// Mitsubishi GX Works2 project: 701125增加出库   PLC: Q10UDEH (continued)
IF iStep=3 AND ConveyorMotor.xSizeDeficientDetect AND (NOT ConveyorMotor.xCCWPresent OR NOT ConveyorMotor.xCWPresent)  THEN
	   ConveyorMotor.xOverWidthAlarm:=1;
	    iStep:=0;               
END_IF;
(*//总报警*)
ConveyorMotor.xError:=ConveyorMotor.xLimitAlarrm
                                              OR ConveyorMotor.xNotArriveAlarm
                                              OR ConveyorMotor.xUnloadAlarm                                             
                                              OR ConveyorMotor.xOverWidthAlarm;

(*//状态输出*)(*状态显示，容易造成指针容量不足*)
IF ConveyorMotor.xEmpty AND NOT ConveyorMotor.xBusy THEN
	m_wStateWord:=0;
END_IF;
IF ConveyorMotor.xEmpty=0 THEN
		m_wStateWord:=1;
END_IF;
IF ConveyorMotor.xBusy THEN
		m_wStateWord:=2;
END_IF;
IF ConveyorMotor.xLimitAlarrm THEN
		m_wStateWord:=3;
END_IF;
IF ConveyorMotor.xOverWidthAlarm THEN
		m_wStateWord:=4;
END_IF;
IF ConveyorMotor.xNotArriveAlarm THEN	
		m_wStateWord:=5;
END_IF;
IF ConveyorMotor.xUnloadAlarm THEN
		m_wStateWord:=6;	
END_IF;
(*选择本线体后，将状态赋值给全局变量进行显示*)
IF ConveyorMotor.iDeviceID=g_iDeviceIDSelect THEN
	g_iConveyorStatus:=m_wStateWord;
END_IF;
END_FUNCTION_BLOCK

FUNCTION_BLOCK DivideFolder
VAR_IN_OUT
  FolderIO : FolderIO;
  FolderConveyorIO : ConveyorIO;
END_VAR
VAR
  iFolderCount : INT;
  m_xInitial : BOOL;
  istep : INT;
  m_TONLoadDelay : TON;  (* 上料完成延时 *)
  m_xLoadDelay : BOOL;  (* 上料完成延时 *)
  m_tLoadDelay : TIME;  (* 上料完成延时 *)
  m_TONUpCylinderError : TON;
  m_tUpCylinderError : TIME;
  m_TONDownCylinderError : TON;
  m_tDownCylinderError : TIME;
  m_TONGrabCylinderError : TON;
  m_tGrabCylinderError : TIME;
END_VAR
VAR_INPUT
  i_xAuto : BOOL;  (* 自动 *)
END_VAR
(*拆盘机*)
(*Mr.Li修改2018.11.19调试*)
(*初始化*)
IF NOT m_xInitial  THEN
	FolderIO.i_iFloor:=3;
	 iFolderCount:=3;
	 	FolderIO.i_tSetOvertime:=T#5S;
		m_xInitial:=1;
END_IF;
(*自动*)
IF i_xAuto THEN
	FolderIO.o_xEntryPermit:=iFolderCount=3 AND FolderConveyorIO.xEmpty;(*线体状态为空且拆盘初始数量为3，才准上料*)
	m_TONLoadDelay(IN:= NOT FolderConveyorIO.xEmpty,
											PT:= T#100MS,
											Q:=m_xLoadDelay,
											ET:=m_tLoadDelay);

	CASE istep OF
		0:(*各种初始化*)
			FolderConveyorIO.xLoad:=0;
			FolderConveyorIO.xUnload:=0;
			FolderConveyorIO.xPutInto:=0;
			IF FolderConveyorIO.xEmpty THEN(*空的情况，0时上料，其他走流程*)
				IF iFolderCount=FolderIO.i_iFloor   THEN
					istep:=1; 					
				ELSE
					istep:=5;
				END_IF;	
			END_IF;		
			IF m_xLoadDelay THEN
				 IF FolderIO.i_xCylinderDownRetractDetect AND FolderIO.i_xCylinderUpRetractDetect THEN
					istep:=2;(*如果在1层，则顶起，需人为判断是否在指定位置，否则有翻框的危险*)
				ELSE
				 	istep:=3;(*如果有料不在1层，则抓紧，然后跳到第4步判断是否是叠盘，不是就放行*)
				 END_IF;
			END_IF;
		1:(*上料*)
			IF FolderIO.o_xEntryPermit THEN
				FolderConveyorIO.xLoad:=FolderIO.i_FrontConveyorNextRun;
			ELSE
				FolderConveyorIO.xLoad:=0;
			END_IF;(*有料等延时*)	
			IF m_xLoadDelay THEN
				iFolderCount:=FolderIO.i_iFloor;
				istep:=2;(**拆盘机顶起步骤*)
			END_IF;	
		2:(*上升至2层位置*)
				FolderIO.o_xCylinderDownRetract:=0;
				FolderIO.o_xCylinderDownExtend:=1;
				FolderIO.o_xCylinderUpRetract:=0;
				IF FolderIO.i_xCylinderDownExtendDetect   THEN
				istep:=3;
				END_IF;
		3:	(*夹紧夹爪*)
			IF FolderIO.i_xCylinderDownExtendDetect THEN
				FolderIO.o_xCylinderGrabExtend:=1;
				FolderIO.o_xCylinderGrabRetract:=0;
			END_IF;
			IF FolderIO.i_xCylinderGrabExtendDetect THEN
				istep:=4;
			END_IF;	
		4:(*再下降到1层，然后放行，在该位置判断是不是最后一次*)
				FolderIO.o_xCylinderUpRetract:=1;
				FolderIO.o_xCylinderUpExtend:=0;
				FolderIO.o_xCylinderDownRetract:=1;
				FolderIO.o_xCylinderDownExtend:=0;
				IF FolderIO.i_xCylinderDownRetractDetect AND FolderIO.i_xCylinderUpRetractDetect AND FolderIO.o_xExitPremit THEN
				FolderConveyorIO.xPutInto:=1;
				FolderConveyorIO.xUnload:=FolderIO.o_xExitPremit;
				ELSIF NOT FolderIO.i_xTrayDetect AND NOT FolderConveyorIO.xEmpty AND FolderIO.o_xExitPremit THEN 
						FolderConveyorIO.xUnload:=FolderIO.o_xExitPremit;
				ELSE 
					FolderConveyorIO.xPutInto:=0;
				FolderConveyorIO.xUnload:=0;
				END_IF;
					IF FolderIO.i_xCylinderDownRetractDetect AND FolderIO.i_xCylinderUpRetractDetect AND
						  FolderIO.i_xTrayDetect  AND  iFolderCount>0  AND ldp(TRUE,NOT  FolderConveyorIO.xUnload) THEN
						iFolderCount:=FolderIO.i_iFloor-1;					
					istep:=5;
					ELSIF  FolderIO.i_xCylinderDownRetractDetect AND FolderIO.i_xCylinderUpRetractDetect  AND 
						 NOT FolderIO.i_xTrayDetect   AND  FolderConveyorIO.xEmpty THEN 
						 	istep:=7;
					END_IF;

		5:(*上升到3层*)
			FolderIO.o_xCylinderUpRetract:=0;
			FolderIO.o_xCylinderUpExtend:=1;
			FolderIO.o_xCylinderDownRetract:=0;
			IF  FolderIO.i_xCylinderUpExtendDetect THEN
				istep:=6;
			END_IF;		
		6:(*松开并下降*)
			FolderIO.i_iFloor:=iFolderCount;
			IF  FolderIO.i_xCylinderUpExtendDetect  THEN
				FolderIO.o_xCylinderGrabExtend:=0;
				FolderIO.o_xCylinderGrabRetract:=1;
				IF FolderIO.i_xCylinderGrabRetractDetect THEN
					FolderIO.o_xCylinderUpRetract:=1;
					FolderIO.o_xCylinderUpExtend:=0;
					FolderIO.o_xCylinderDownRetract:=1;
					FolderIO.o_xCylinderDownExtend:=0;
				END_IF;		
			END_IF;	
			IF   FolderIO.i_xCylinderUpRetractDetect  AND FolderIO.i_xCylinderDownRetractDetect  THEN
				istep:=2;
			ELSIF iFolderCount=0 THEN 
				istep:=7;
			ELSIF  NOT FolderIO.i_xTrayDetect  THEN 
				istep:=4;
			END_IF;	
			
		7:(*恢复初始状态*)	
			FolderIO.o_xCylinderDownRetract:=1;
			FolderIO.o_xCylinderUpRetract:=1;
			FolderIO.o_xCylinderDownExtend:=0;
			FolderIO.o_xCylinderUpExtend:=0;
			FolderIO.o_xCylinderGrabExtend:=0;
			FolderIO.o_xCylinderGrabRetract:=1;
			iFolderCount:=3;
			FolderIO.i_iFloor:=3;
			IF FolderIO.i_xCylinderDownRetractDetect  AND FolderIO.i_xCylinderUpRetractDetect THEN 
			istep:=0;
			END_IF;
		END_CASE;
END_IF;(*g_xAuto那个*)	
(*手动控制气缸动作*)
		IF NOT i_xAuto THEN
			FolderIO.o_xCylinderGrabExtend:=	FolderIO.i_xCylinderGrabExtendButton;	
			FolderIO.o_xCylinderGrabRetract:=	FolderIO.i_xCylinderGrabRetractButton;	
			FolderIO.o_xCylinderUpExtend:=		FolderIO.i_xCylinderUpExtendButton;	
			FolderIO.o_xCylinderUpRetract:=		FolderIO.i_xCylinderUpRetractButton;	
			FolderIO.o_xCylinderDownExtend:=	FolderIO.i_xCylinderDownExtendButton;	
			FolderIO.o_xCylinderDownRetract:=	FolderIO.i_xCylinderDownRetractButton;		
		END_IF;
		
		(*气缸超时未到达报警，可能是没气儿漏气，也可能是开关坏了，或者气缸被卡住了*)
		m_TONGrabCylinderError(IN:= (FolderIO.o_xCylinderGrabExtend AND NOT FolderIO.i_xCylinderGrabExtendDetect) 
																OR  (FolderIO.o_xCylinderGrabRetract AND NOT FolderIO.i_xCylinderGrabRetractDetect) ,
															PT:= FolderIO.i_tSetOvertime ,Q:= FolderIO.o_xGrabCylinderError,ET:= m_tGrabCylinderError);
		m_TONDownCylinderError(IN:= (FolderIO.o_xCylinderDownExtend AND NOT FolderIO.i_xCylinderDownExtendDetect) 
																OR  (FolderIO.o_xCylinderDownRetract AND NOT FolderIO.i_xCylinderDownRetractDetect) ,
															PT:= FolderIO.i_tSetOvertime ,Q:= FolderIO.o_xDownCylinderError,ET:= m_tDownCylinderError);
		m_TONUpCylinderError(IN:= (FolderIO.o_xCylinderUpExtend AND NOT FolderIO.i_xCylinderUpExtendDetect) 
																OR  (FolderIO.o_xCylinderUpRetract AND NOT FolderIO.i_xCylinderUpRetractDetect) ,
															PT:= FolderIO.i_tSetOvertime ,Q:= FolderIO.o_xUpCylinderError,ET:= m_tUpCylinderError);
END_FUNCTION_BLOCK

FUNCTION_BLOCK FanucRobot
VAR_IN_OUT
  FanucRobotIO : FanucRobotIO;
END_VAR
VAR
  m_iSNO : INT;
  m_xPNSPass : BOOL;  (* 收到程序号 *)
  m_tonStartDelay : TON;  (* 启动延时 *)
  m_xStartDelay : BOOL;
  m_tStartDelayCurrentTime : TIME;
END_VAR
(***********************************************************
发那科机器人自动启动程序


***********************************************************)

(*无自动状态，示教盒处于本地状态，把各标志位复位*)
IF FanucRobotIO.i_xTPENBL AND NOT g_xAuto THEN
	FanucRobotIO.o_xPNSTROBE:=0;
	FanucRobotIO.o_xCSTOPI:=0;
	FanucRobotIO.o_xPROD_START:=0;
	FanucRobotIO.o_xRESET:=0;
END_IF;
(*远程模式*)
IF g_xAuto THEN
	FanucRobotIO.o_xREMOTE:=1;
	ELSE
	FanucRobotIO.o_xREMOTE:=0;
END_IF;
(*程序启动后复位启动标志位*)
IF FanucRobotIO.i_xPROG_RUN AND FanucRobotIO.i_xBUSY THEN
	FanucRobotIO.i_xCommandStart:=0;
END_IF;
(*示教盒旋清除报警*)
IF ldf(TRUE,FanucRobotIO.i_xTPENBL)THEN
	FanucRobotIO.o_xRESET:=1;
	FanucRobotIO.o_xCSTOPI:=1;
END_IF;
(*启动程序号条件*)
IF FanucRobotIO.i_xSYSRDY 
	AND FanucRobotIO.i_xCMDENBL
	AND FanucRobotIO.i_xCommandStart
	AND NOT FanucRobotIO.i_xPROG_RUN 
	AND NOT FanucRobotIO.i_xBUSY THEN
	FanucRobotIO.o_xRESET:=0;
	FanucRobotIO.o_xCSTOPI:=0;
	IF FanucRobotIO.i_iMotionNumber <> 0 (*只要动作编号不为0，就给他信号*)
		AND NOT FanucRobotIO.o_xPNSTROBE THEN
		FanucRobotIO.o_xPNSTROBE:=1;
		FanucRobotIO.o_xPROD_START:=1;
		FanucRobotIO.o_iPNS:=FanucRobotIO.i_iMotionNumber;(*并把任务号传给他*)
	END_IF;
	(*程序号校验*)
	IF FanucRobotIO.i_xSNACK THEN(*数据传回之后再校验*)
		m_iSNO:=BITARR_TO_INT(FanucRobotIO.i_arrxSNO[0] , 8 );
		IF m_iSNO=FanucRobotIO.o_iPNS THEN
			m_xPNSPass:=1;(*校验成功,等100MS复位Start信号*)
			FanucRobotIO.o_xPNSTROBE:=0;
		ELSE
			FanucRobotIO.o_xPNSFailed:=1;(*校验失败*)
			FanucRobotIO.o_xPROD_START:=0;(*立刻复位，不生成任务*)
		END_IF;
	END_IF;
END_IF;
m_tonStartDelay(IN:= m_xPNSPass ,PT:= T#100ms ,Q:= m_xStartDelay ,ET:=m_tStartDelayCurrentTime );
IF m_xStartDelay THEN
	FanucRobotIO.o_xPROD_START:=0;
	FanucRobotIO.i_xCommandStart:=0;
	m_xPNSPass:=0;
END_IF;
END_FUNCTION_BLOCK

FUNCTION_BLOCK Folder
VAR_IN_OUT
  FolderIO : FolderIO;
END_VAR
VAR
  m_xInitial : BOOL;
END_VAR
VAR_IN_OUT
  FolderConveyorIO : ConveyorIO;
END_VAR
VAR
  iFolderCount : INT;
  istep : INT;
  m_TONLoadDelay : TON;  (* 上料完成延时 *)
  m_xLoadDelay : BOOL;  (* 上料完成延时 *)
  m_tLoadDelay : TIME;  (* 上料完成延时 *)
  m_TONUpCylinderError : TON;
  m_tUpCylinderError : TIME;
  m_TONDownCylinderError : TON;
  m_tDownCylinderError : TIME;
  m_TONGrabCylinderError : TON;
  m_tGrabCylinderError : TIME;
END_VAR
VAR_INPUT
  i_xAuto : BOOL;  (* 自动 *)
  i_xManual : BOOL;  (* 手动 *)
END_VAR
(*叠盘机*)
(*sb刘写的*)
(*初始化*)
(*18/11/17 YAOBO更改*)
(*增加允许下料信号o_xExitPrimit，码垛完成后给允许下料第7步给出*)
IF NOT m_xInitial THEN
	FolderIO.i_iFloor:=3;
	FolderIO.i_tSetOvertime:=T#5S;
	
	m_xInitial:=1;
END_IF;
(*自动*)
FolderIO.o_xEntryPermit:=FolderConveyorIO.xEmpty;(*叠盘机的话，只要空了，就允许上料，拆盘则是拆完才允许*)
IF i_xAuto THEN
				m_TONLoadDelay(IN:= NOT FolderConveyorIO.xEmpty,
													PT:= T#100MS,
													Q:=m_xLoadDelay,
													ET:=m_tLoadDelay);
	CASE istep OF
		0:(*各种初始化*)
			FolderConveyorIO.xLoad:=0;
			FolderConveyorIO.xUnload:=0;
			FolderConveyorIO.xPutInto:=0;
			FolderIo.o_xExitPremit:=0;	
			IF (*0 AND*)  FolderConveyorIO.xEmpty THEN
				istep:=1;(*空着就去1上料*)
			END_IF;	
			IF 0 AND    m_xLoadDelay  THEN(*if 有料*)
				IF  FolderIO.i_xCylinderDownExtendDetect  AND FolderIO.i_xCylinderUpExtendDetect  THEN(*if 在下层*)
					IF iFolderCount=FolderIO.i_iFloor THEN(*if 是最后一次*)
						istep:=7;
					ELSE(*不是最后一次去5，是就去7*)
						istep:=5;
					END_IF;(*if 是最后一次*)	
				ELSE(*不在下层去2*)
				istep:=2;
				END_IF;	(*if 在下层*)			
			END_IF;(*if 有料*)
			
		1:(*上料*)
			IF FolderIO.i_xEntryEnable THEN
				FolderConveyorIO.xLoad:=1;
			ELSE
				FolderConveyorIO.xLoad:=0;
			END_IF;(*not Empty了等个延时*)	

			IF (*0 AND*)   m_xLoadDelay  AND (iFolderCount>0 AND iFolderCount<FolderIO.i_iFloor) THEN
				istep:=2;
			ELSIF (*0 AND*)   m_xLoadDelay AND iFolderCount=0 THEN(*=0表示是第一次，第一次直接抓紧上升*)
				istep:=5;	
			END_IF;	
		2:(*下降，到2层位置*)
				FolderIO.o_xCylinderUpRetract:=0;
				FolderIO.o_xCylinderUpExtend:=1;
				FolderIO.o_xCylinderDownRetract:=1;
				FolderIO.o_xCylinderDownExtend:=0;
				IF FolderIO.i_xCylinderUpExtendDetect AND NOT FolderIO.i_xCylinderDownExtendDetect THEN
					istep:=3;
				END_IF;
		3:	(*松开夹爪*)
			IF FolderConveyorIO.xCWPresent AND NOT FolderConveyorIO.xEmpty THEN(*有感应到才松开*)
				FolderIO.o_xCylinderGrabExtend:=0;
				FolderIO.o_xCylinderGrabRetract:=1;
				IF (*0 AND*)   FolderIO.i_xCylinderGrabRetractDetect THEN
					IF iFolderCount=FolderIO.i_iFloor-1 THEN
						iFolderCount:=FolderIO.i_iFloor;(*最后一次到这里就刷新计数，方便故障恢复*)
					END_IF;	
					istep:=4;
				END_IF;	
			END_IF;	
		4:(*再下降，去1层*)
				FolderIO.o_xCylinderUpRetract:=0;
				FolderIO.o_xCylinderUpExtend:=1;
				FolderIO.o_xCylinderDownRetract:=0;
				FolderIO.o_xCylinderDownExtend:=1;
				IF FolderIO.i_xCylinderDownExtendDetect  AND FolderIO.i_xCylinderUpExtendDetect  THEN
					IF iFolderCount<FolderIO.i_iFloor-1 THEN
						istep:=5;
					ELSE
						istep:=7;
					END_IF;	
				END_IF;		
		5:(*抓紧*)
			IF FolderIO.i_xCylinderDownExtendDetect  AND FolderIO.i_xCylinderUpExtendDetect  THEN
				FolderIO.o_xCylinderGrabExtend:=1;
				FolderIO.o_xCylinderGrabRetract:=0;
				IF (*0 AND*)   FolderIO.i_xCylinderGrabExtendDetect THEN
					iFolderCount:=iFolderCount+1;
					istep:=6;
				END_IF;	
			END_IF;		
		6:(*上升到3层*)
			FolderIO.o_xCylinderUpRetract:=1;
			FolderIO.o_xCylinderUpExtend:=0;
			FolderIO.o_xCylinderDownRetract:=1;
			FolderIO.o_xCylinderDownExtend:=0;
			IF (*0 AND *)  FolderIO.i_xCylinderDownRetractDetect AND FolderIO.i_xCylinderUpRetractDetect THEN
				FolderConveyorIO.xPutInto:=1;(*刷新成Empty的*)
				istep:=0;
			END_IF;
		7:(*下料*)
		FolderIo.o_xExitPremit:=1;	(*给出允许下料信号*)
		FolderConveyorIO.xUnload:=	FolderIO.i_xExitEnable AND FolderIO.i_xCylinderGrabRetractDetect;(*给下料信号，不要刷新完成*)
	(*			IF	FolderIO.i_xExitEnable AND FolderIO.i_xCylinderGrabRetractDetect	THEN(*保证不会挂到叉手*)
(*				FolderConveyorIO.xUnload:=1;
			ELSE
				FolderConveyorIO.xPutInto:=1;(*刷新成Empty的*)
	(*			FolderConveyorIO.xUnload:=0;
			END_IF;	*)
			IF FolderConveyorIO.xEmpty THEN(*确保空了才回0，不然还在这里等Unload信号*)
				iFolderCount:=0;
				istep:=0;
			END_IF;	 
		END_CASE;
END_IF;(*g_xAuto那个*)	
(*手动控制气缸动作*)
		IF i_xManual THEN
			FolderIO.o_xCylinderGrabExtend:=	FolderIO.i_xCylinderGrabExtendButton;	
			FolderIO.o_xCylinderGrabRetract:=	FolderIO.i_xCylinderGrabRetractButton;	
			FolderIO.o_xCylinderUpExtend:=		FolderIO.i_xCylinderUpExtendButton;	
			FolderIO.o_xCylinderUpRetract:=		FolderIO.i_xCylinderUpRetractButton;	
			FolderIO.o_xCylinderDownExtend:=	FolderIO.i_xCylinderDownExtendButton;	
			FolderIO.o_xCylinderDownRetract:=	FolderIO.i_xCylinderDownRetractButton;		
		END_IF;
		
		(*气缸超时未到达报警，可能是没气儿漏气，也可能是开关坏了，或者气缸被卡住了*)
		m_TONGrabCylinderError(IN:= (FolderIO.o_xCylinderGrabExtend AND NOT FolderIO.i_xCylinderGrabExtendDetect) 
																OR  (FolderIO.o_xCylinderGrabRetract AND NOT FolderIO.i_xCylinderGrabRetractDetect) ,
															PT:= FolderIO.i_tSetOvertime ,Q:= FolderIO.o_xGrabCylinderError,ET:= m_tGrabCylinderError);
		m_TONDownCylinderError(IN:= (FolderIO.o_xCylinderDownExtend AND NOT FolderIO.i_xCylinderDownExtendDetect) 
																OR  (FolderIO.o_xCylinderDownRetract AND NOT FolderIO.i_xCylinderDownRetractDetect) ,
															PT:= FolderIO.i_tSetOvertime ,Q:= FolderIO.o_xDownCylinderError,ET:= m_tDownCylinderError);
		m_TONUpCylinderError(IN:= (FolderIO.o_xCylinderUpExtend AND NOT FolderIO.i_xCylinderUpExtendDetect) 
																OR  (FolderIO.o_xCylinderUpRetract AND NOT FolderIO.i_xCylinderUpRetractDetect) ,
															PT:= FolderIO.i_tSetOvertime ,Q:= FolderIO.o_xUpCylinderError,ET:= m_tUpCylinderError);
END_FUNCTION_BLOCK

FUNCTION_BLOCK FolderII
VAR_IN_OUT
  FolderIO : FolderIO;
  FolderConveyorIO : ConveyorIO;
END_VAR
VAR_INPUT
  i_xAuto : BOOL;  (* 自动 *)
END_VAR
VAR
  iFolderCount : INT;
  m_xInitial : BOOL;
  istep : INT;
  m_TONLoadDelay : TON;  (* 上料完成延时 *)
  m_xLoadDelay : BOOL;  (* 上料完成延时 *)
  m_tLoadDelay : TIME;  (* 上料完成延时 *)
  m_TONUpCylinderError : TON;
  m_tUpCylinderError : TIME;
  m_TONDownCylinderError : TON;
  m_tDownCylinderError : TIME;
  m_TONGrabCylinderError : TON;
  m_tGrabCylinderError : TIME;
END_VAR
VAR_INPUT
  i_xManual : BOOL;  (* 手动 *)
END_VAR
(*叠盘机II型*)
(*初始化*)
(*18/11/17 YAOBO更改*)
(*增加允许下料信号o_xExitPrimit，码垛完成后给允许下料第7步给出*)
IF NOT m_xInitial THEN
	FolderIO.i_iFloor:=3;
	FolderIO.i_tSetOvertime:=T#5S;
	
	m_xInitial:=1;
END_IF;
(*自动*)
FolderIO.o_xEntryPermit:=FolderConveyorIO.xEmpty;(*叠盘机的话，只要空了，就允许上料，拆盘则是拆完才允许*)
IF i_xAuto THEN
				m_TONLoadDelay(IN:= NOT FolderConveyorIO.xEmpty,
													PT:= T#100MS,
													Q:=m_xLoadDelay,
													ET:=m_tLoadDelay);
	CASE istep OF
		0:(*各种初始化*)
			FolderConveyorIO.xLoad:=0;
			FolderConveyorIO.xUnload:=0;
			FolderConveyorIO.xPutInto:=0;
			FolderIo.o_xExitPremit:=0;	
			FolderIo.i_xExitEnable:=0;
			IF (*0 AND*)  FolderConveyorIO.xEmpty THEN
				istep:=1;(*空着就去1上料*)
			END_IF;	
			IF 0 AND    m_xLoadDelay  THEN(*if 有料*)
				IF  FolderIO.i_xCylinderDownRetractDetect  AND FolderIO.i_xCylinderUpRetractDetect  THEN(*if 在下层*)
					IF iFolderCount=FolderIO.i_iFloor THEN(*if 是最后一次*)
						istep:=7;
					ELSE(*不是最后一次去5，是就去7*)
						istep:=5;
					END_IF;(*if 是最后一次*)	
				ELSE(*不在下层去2*)
				istep:=2;
				END_IF;	(*if 在下层*)			
			END_IF;(*if 有料*)
			
		1:(*上料*)
			IF FolderIO.i_xEntryEnable THEN
				FolderConveyorIO.xLoad:=1;
			ELSE
				FolderConveyorIO.xLoad:=0;
			END_IF;(*not Empty了等个延时*)	

			IF (*0 AND*)   m_xLoadDelay  AND (iFolderCount>0 AND iFolderCount<FolderIO.i_iFloor) THEN
				istep:=2;
			ELSIF (*0 AND*)   m_xLoadDelay AND iFolderCount=0 THEN(*=0表示是第一次，第一次直接抓紧上升*)
				istep:=4;	
			END_IF;	
		2:(*上升，到2层位置*)
				FolderIO.o_xCylinderUpRetract:=0;
				FolderIO.o_xCylinderUpExtend:=0;
				FolderIO.o_xCylinderDownRetract:=0;
				FolderIO.o_xCylinderDownExtend:=1;
				IF   FolderIO.i_xCylinderDownExtendDetect THEN
					istep:=3;
				END_IF;
		3:	(*松开夹爪,并降到1层*)
			IF  FolderIO.i_xTrayDetect AND NOT FolderConveyorIO.xEmpty THEN(*有感应到才松开*)
				FolderIO.o_xCylinderGrabExtend:=0;
				FolderIO.o_xCylinderGrabRetract:=1;
				IF (*0 AND*)   FolderIO.i_xCylinderGrabRetractDetect THEN
					FolderIO.o_xCylinderDownRetract:=1;
					FolderIO.o_xCylinderDownExtend:=0;
					IF iFolderCount=FolderIO.i_iFloor-1 THEN
						iFolderCount:=FolderIO.i_iFloor;(*最后一次到这里就刷新计数，方便故障恢复*)
					END_IF;	
					IF FolderIO.i_xCylinderDownRetractDetect  THEN 
					istep:=4;
					END_IF;
				END_IF;	
			END_IF;	
		4:(*再上升，去3层*)
		IF iFolderCount<FolderIO.i_iFloor-1 THEN 
				FolderIO.o_xCylinderUpRetract:=0;
				FolderIO.o_xCylinderUpExtend:=1;
				FolderIO.o_xCylinderDownRetract:=0;
				FolderIO.o_xCylinderDownExtend:=0;
				IF  FolderIO.i_xCylinderUpExtendDetect
					THEN  istep:=5;
				END_IF;
		ELSE FolderIO.o_xCylinderUpRetract:=1;
				FolderIO.o_xCylinderUpExtend:=0;
				FolderIO.o_xCylinderDownRetract:=1;
				FolderIO.o_xCylinderDownExtend:=0;
				   IF  FolderIO.i_xCylinderUpRetractDetect AND FolderIO.i_xCylinderDownRetractDetect THEN 
				   	 istep:=7;
				   END_IF;
		END_IF;
			
	
		5:(*抓紧*)
			IF  FolderIO.i_xCylinderUpExtendDetect  THEN
				FolderIO.o_xCylinderGrabExtend:=1;
				FolderIO.o_xCylinderGrabRetract:=0;
				IF (*0 AND*)   FolderIO.i_xCylinderGrabExtendDetect THEN
					iFolderCount:=iFolderCount+1;
					istep:=6;
				END_IF;	
			END_IF;		
		6:(*下降到1层*)
			FolderIO.o_xCylinderUpRetract:=1;
			FolderIO.o_xCylinderUpExtend:=0;
			FolderIO.o_xCylinderDownRetract:=1;
			FolderIO.o_xCylinderDownExtend:=0;
			IF (*0 AND *)  FolderIO.i_xCylinderDownRetractDetect AND FolderIO.i_xCylinderUpRetractDetect THEN
				FolderConveyorIO.xPutInto:=1;(*刷新成Empty的*)
				istep:=0;
			END_IF;
		7:(*下料*)
		FolderIo.o_xExitPremit:=1;	(*给出允许下料信号*)
		IF FolderIo.o_xExitPremit
			THEN FolderIo.i_xExitEnable:=1;
		END_IF;
		FolderConveyorIO.xUnload:=	FolderIO.i_NextConveyorEmpty AND FolderIO.i_xCylinderGrabRetractDetect AND
		 FolderIO.i_xCylinderDownRetractDetect AND FolderIO.i_xCylinderUpRetractDetect ;(*给下料信号，不要刷新完成*)
	(*			IF	FolderIO.i_xExitEnable AND FolderIO.i_xCylinderGrabRetractDetect	THEN(*保证不会挂到叉手*)
(*				FolderConveyorIO.xUnload:=1;
			ELSE
				FolderConveyorIO.xPutInto:=1;(*刷新成Empty的*)
	(*			FolderConveyorIO.xUnload:=0;
			END_IF;	*)
			IF FolderConveyorIO.xEmpty THEN(*确保空了才回0，不然还在这里等Unload信号*)
				iFolderCount:=0;
				istep:=0;
			END_IF;	 
		END_CASE;
END_IF;(*g_xAuto那个*)	
(*手动控制气缸动作*)
		IF i_xManual THEN
			FolderIO.o_xCylinderGrabExtend:=	FolderIO.i_xCylinderGrabExtendButton;	
			FolderIO.o_xCylinderGrabRetract:=	FolderIO.i_xCylinderGrabRetractButton;	
			FolderIO.o_xCylinderUpExtend:=		FolderIO.i_xCylinderUpExtendButton;	
			FolderIO.o_xCylinderUpRetract:=		FolderIO.i_xCylinderUpRetractButton;	
			FolderIO.o_xCylinderDownExtend:=	FolderIO.i_xCylinderDownExtendButton;	
			FolderIO.o_xCylinderDownRetract:=	FolderIO.i_xCylinderDownRetractButton;		
		END_IF;
		
		(*气缸超时未到达报警，可能是没气儿漏气，也可能是开关坏了，或者气缸被卡住了*)
		m_TONGrabCylinderError(IN:= (FolderIO.o_xCylinderGrabExtend AND NOT FolderIO.i_xCylinderGrabExtendDetect) 
																OR  (FolderIO.o_xCylinderGrabRetract AND NOT FolderIO.i_xCylinderGrabRetractDetect) ,
															PT:= FolderIO.i_tSetOvertime ,Q:= FolderIO.o_xGrabCylinderError,ET:= m_tGrabCylinderError);
		m_TONDownCylinderError(IN:= (FolderIO.o_xCylinderDownExtend AND NOT FolderIO.i_xCylinderDownExtendDetect) 
																OR  (FolderIO.o_xCylinderDownRetract AND NOT FolderIO.i_xCylinderDownRetractDetect) ,
															PT:= FolderIO.i_tSetOvertime ,Q:= FolderIO.o_xDownCylinderError,ET:= m_tDownCylinderError);
		m_TONUpCylinderError(IN:= (FolderIO.o_xCylinderUpExtend AND NOT FolderIO.i_xCylinderUpExtendDetect) 
																OR  (FolderIO.o_xCylinderUpRetract AND NOT FolderIO.i_xCylinderUpRetractDetect) ,
															PT:= FolderIO.i_tSetOvertime ,Q:= FolderIO.o_xUpCylinderError,ET:= m_tUpCylinderError);
END_FUNCTION_BLOCK

FUNCTION_BLOCK PackCommunication
VAR_IN_OUT
  ConveyorIO : ConveyorIO;
  PackCommunicationIO : PackCommunicationIO;
  FanucRobotIO : FanucRobotIO;
END_VAR
VAR_OUTPUT
  o_iErrorNub : INT;
  o_xReqSuccess : BOOL;
END_VAR
VAR
  m_xReqSuccess : BOOL;
  m_iStep : INT;
  m_arrwCode : ARRAY [1..8] OF BatteryCode;
END_VAR
VAR_INPUT
  i_arrxPresentDetect : ARRAY [1..8] OF BOOL;
END_VAR
VAR
  m_iCoordinateX : INT;
  m_iCoordinateY : INT;
  m_arriPresentDetect : ARRAY [1..8] OF INT;
  ii : INT;
END_VAR
VAR CONSTANT
  MAX_ROW : INT := 8;
  MAX_COLUMN : INT := 8;
END_VAR
VAR
  m_xSupplement : BOOL;
END_VAR
VAR CONSTANT
  ROW_TIMES : INT := 1;
  GET_QUANTITY : INT := 8;
END_VAR
VAR
  m_iRowReminder : INT;
  m_xEno : BOOL;
  m_iRowReminderTemp : INT;
END_VAR
(***************************************************************************)
(*
DB1区(PC->PLC)10个字		
"字(16位）序号
(从1开始)"	功能描述	具体参数解释
1	请求确认	"1：复位
2：读码(入库申请）成功
101：条码空
102：条码规则校验失败
103：步号校验失败
"
2	放行	"1：复位
2：完成,放行
3：撤销完成 "
3	单次装载应答	"1：复位
2：允许开始"
4	单次装载处理完成	"1：复位
2：完成
3：电芯为空"
)*
DB2区(PLC->PC)200个字		
"字(16位）序号
(从1开始)"	功能描述	具体参数解释
1	装载请求	"１：复位
２：请求"
2	装载全部完成	"1：复位
2：请求 "
3	单次装载请求	"1：复位
2：请求 "
4	单次装载完成	"1：复位
2：完成"
5	行坐标	从1开始
6	列坐标	从1开始
7	电芯码(15*11=165)	"电芯码24字符，
占12个字，加上预留的每个分配15个字"

顺序执行步骤
0  初始化
1  框码扫码请求
2  单次抓取请求
3  整排抓取
4  补料
5  完成


(***************************************************************************)
m_iRowReminder:= ( m_iCoordinateX-1 MOD GET_QUANTITY )+1;(*//通过位置与抓取数量取余数，判断是否的抓取位置为一排的最后一个*)
CASE m_iStep OF
	0:;(*//初始化*)
	m_iStep:=1;
	1:(*发送框码的扫码请求*)
	IF NOT ConveyorIO.xEmpty AND NOT FanucRobotIO.io_xMutexLock THEN
		PackCommunicationIO.o_iRequestPLCPC:=2;
		ELSE
		PackCommunicationIO.o_iRequestPLCPC:=1;
	END_IF;
	(*//请求确认*)
	CASE PackCommunicationIO.i_iResponsPCPLC OF 
		0:;
		1:;(*//复位*)
		2:(*//读码（入库申请）成功*)
		m_iStep:=2;
		m_xSupplement:=0;
		m_iCoordinateX:=1;(*//框码扫码成功后把坐标改为1,1*)
		m_iCoordinateY:=1;
		FanucRobotIO.io_xMutexLock:=1;
		3:(*//取放货完成*)
		ConveyorIO.xPutInto:=1; 
		4:(*//旋转*)
		;
		5:(*//不旋转*)
		;
		101:(*//条码空*)
		o_iErrorNub:=101;
		m_iStep:=0;
		102:(*//条码规则检验失败*)
		o_iErrorNub:=102;
		m_iStep:=0;
		103:(*//步号校验失败*)
		o_iErrorNub:=103;
		m_iStep:=0;
		104:(*//无库位可用*)
		o_iErrorNub:=104;
		m_iStep:=0;
	END_CASE;
	2:(*//单次抓取请求，分为单次多个产品抓取与补料程序*)
	IF FanucRobotIO.i_xSYSRDY 
		AND NOT FanucRobotIO.i_xBUSY
		AND NOT FanucRobotIO.i_xPROG_RUN
		AND i_arrxPresentDetect[1] 
		AND PackCommunicationIO.i_iSinglePackResponsePCPLC=1 THEN(*//机器人准备就绪、组装下线有料*)
		PackCommunicationIO.o_iSinglePackRequestPLCPC:=2;
	END_IF;
	IF (*LDP(TRUE,PackCommunicationIO.i_iSinglePackResponsePCPLC=2)*) PackCommunicationIO.i_iSinglePackResponsePCPLC=2 THEN(*//请求成功*)
		PackCommunicationIO.o_iSinglePackRequestPLCPC:=1;(*//复位请求*)
		IF m_xSupplement THEN(*//补料标志位，为1进行补料操作，为0进行整排抓取*)
			m_iStep:=4;(*//补料*)
			ELSE
		 	m_iStep:=3;(*//整排抓取*)
			FOR ii:=1 TO GET_QUANTITY BY 1 DO(*//记录哪个位置缺料*)
				IF i_arrxPresentDetect[ii] THEN(*//传感器检测*)
 m_arriPresentDetect[ii]:=0;
 ELSE
 m_arriPresentDetect[ii]:=ii;(*//记录缺料的位置*)
				END_IF;
			END_FOR;
		END_IF;
	END_IF;
	3:  (*//整排抓取*)
	FanucRobotIO.o_iPNS:=10101;(*//步骤号*)
	FanucRobotIO.o_uiOffset_X:=m_iCoordinateX;
	FanucRobotIO.o_uiOffset_Y:=m_iCoordinateY;
	PackCommunicationIO.o_iXCoordinatePLCPC:=m_iCoordinateX;(*//放置位置发送给上位机*)
	PackCommunicationIO.o_iYCoordinatePLCPC:=m_iCoordinateY;	
	IF LDF(TRUE,FanucRobotIO.i_xBUSY OR FanucRobotIO.i_xPROG_RUN) THEN(*//抓取动作完成*)
		FOR ii:=1 TO GET_QUANTITY BY 1 DO (*//判断有无补料信息*)
			IF m_arriPresentDetect[ii]<>0  THEN(*//有补料*)(*//补料不是最后一个的算法*)
				m_iCoordinateX:=m_arriPresentDetect[ii]+((m_iCoordinateX-1)/GET_QUANTITY)*GET_QUANTITY;
				m_xSupplement:=1;
				m_iStep:=2;(*//有补料*)
				EXIT;
			END_IF;			
		END_FOR;
		IF ii=GET_QUANTITY+1  THEN  (*//无补料*)
			m_xSupplement:=0;
			IF m_iCoordinateY = MAX_ROW (*//达到最大列*)
				AND ((m_iCoordinateX-1)/GET_QUANTITY+1=ROW_TIMES) 
				THEN(*//偏移量为最大的值时,排抓取为最后一排*)
				m_iStep:=5;(*//装盘完成*)
				ELSE
				m_iStep:=2;(*//请求下一次装盘*)			
				IF (m_iCoordinateX-1)/GET_QUANTITY+1=ROW_TIMES THEN
 m_iCoordinateX:=1;                                              (*//开始执行下一列*)
 m_iCoordinateY:=m_iCoordinateY+1;
 ELSE
 m_iCoordinateX:=((m_iCoordinateX-1)/GET_QUANTITY+1)*GET_QUANTITY+1;
				END_IF;
			END_IF;
		END_IF;
	END_IF;
	4: (*//补料*)
	FanucRobotIO.o_iPNS:=10102;(*//步骤号*)
	FanucRobotIO.o_uiOffset_X:=m_iCoordinateX;
	FanucRobotIO.o_uiOffset_Y:=m_iCoordinateY;
	PackCommunicationIO.o_iXCoordinatePLCPC:=m_iCoordinateX;(*//放置位置发送给上位机*)
	PackCommunicationIO.o_iYCoordinatePLCPC:=m_iCoordinateY;
	IF LDF(TRUE,FanucRobotIO.i_xBUSY OR FanucRobotIO.i_xPROG_RUN) THEN(*//抓取动作完成*)
		FOR ii:=m_iRowReminder+1 TO GET_QUANTITY BY 1 DO (*//判断有无补料信息*)
			IF m_arriPresentDetect[ii]<>0  THEN(*//有补料*)(*//补料不是最后一个的算法*)
				m_iCoordinateX:=m_arriPresentDetect[ii]+((m_iCoordinateX-1)/GET_QUANTITY)*GET_QUANTITY;
				m_xSupplement:=1;
				m_iStep:=2;(*//有补料*)
				EXIT;
			END_IF;	
		END_FOR;
		IF ii=GET_QUANTITY+1  THEN  (*//无补料*)
			m_xSupplement:=0;
			IF m_iCoordinateY = MAX_ROW (*//达到最大列*)
				AND ((m_iCoordinateX-1)/GET_QUANTITY+1=ROW_TIMES)
				THEN(*//偏移量为最大的值时,排抓取为最后一排*)
				m_iStep:=5;(*//装盘完成*)
				ELSE
				m_iStep:=2;(*//请求下一次装盘*)			
				IF (m_iCoordinateX-1)/GET_QUANTITY+1=ROW_TIMES THEN
 m_iCoordinateX:=1;                                              (*//开始执行下一列*)
 m_iCoordinateY:=m_iCoordinateY+1;
 ELSE
 m_iCoordinateX:=((m_iCoordinateX-1)/GET_QUANTITY+1)*GET_QUANTITY+1;(*//这一列继续往后排*)
				END_IF;
			END_IF;
		END_IF;
	END_IF;
	5: (*//完成*)
	PackCommunicationIO.o_iSinglePackDonePLCPC:=2;
	IF PackCommunicationIO.i_iSinglePackDoneAknPCPLC =2 THEN
		PackCommunicationIO.o_iSinglePackDonePLCPC:=1;
		m_iCoordinateX:=1;
		m_iCoordinateY:=1;
		FanucRobotIO.io_xMutexLock:=0;
	END_IF;
	IF ConveyorIO.xEmpty AND PackCommunicationIO.o_iSinglePackDonePLCPC=1 THEN
		m_iStep:=1;
	END_IF;
END_CASE;
END_FUNCTION_BLOCK

PROGRAM POU
VAR
  Conveyor70101 : Conveyor;
  Conveyor70102 : Conveyor;
  Conveyor70103 : Conveyor;
  Conveyor70104 : Conveyor;
  Conveyor70105 : Conveyor;
  Conveyor70106 : Conveyor;
  Conveyor70107 : Conveyor;
  Conveyor70108 : Conveyor;
  Conveyor70109 : Conveyor;
  Conveyor70110 : Conveyor;
  Conveyor70111 : Conveyor;
  Conveyor70112 : Conveyor;
  Conveyor70113 : Conveyor;
  Conveyor70114 : Conveyor;
  Conveyor70115 : Conveyor;
  Conveyor70116 : Conveyor;
  Conveyor70117 : Conveyor;
  Conveyor70118 : Conveyor;
  Conveyor70119 : Conveyor;
  Conveyor70120 : Conveyor;
  Conveyor70121 : Conveyor;
  Conveyor70122 : Conveyor;
  Conveyor70123 : Conveyor;
  Conveyor70124 : Conveyor;
  Conveyor70125 : Conveyor;
  Conveyor70126 : Conveyor;
  Conveyor70127 : Conveyor;
  Conveyor70128 : Conveyor;
  Conveyor70129 : Conveyor;
  Conveyor70130 : Conveyor;
  Conveyor70131 : Conveyor;
  Conveyor70132 : Conveyor;
  Conveyor70133 : Conveyor;
  Conveyor70134 : Conveyor;
  Conveyor70135 : Conveyor;
  Conveyor70136 : Conveyor;
  Conveyor70137 : Conveyor;
  Conveyor70138 : Conveyor;
  Conveyor70139 : Conveyor;
  Conveyor70140 : Conveyor;
  Conveyor70141 : Conveyor;
  Conveyor70142 : Conveyor;
  Conveyor70143 : Conveyor;
  Conveyor70144 : Conveyor;
  Conveyor70145 : Conveyor;
  Conveyor70146 : Conveyor;
  Conveyor70147 : Conveyor;
  Conveyor70148 : Conveyor;
  Conveyor70149 : Conveyor;
  Conveyor70150 : Conveyor;
  Conveyor70151 : Conveyor;
  Conveyor70152 : Conveyor;
  Conveyor70153 : Conveyor;
  Conveyor70154 : Conveyor;
  Conveyor70155 : Conveyor;
  Conveyor70156 : Conveyor;
  Conveyor70157 : Conveyor;
  Conveyor70158 : Conveyor;
  Conveyor70159 : Conveyor;
  Conveyor70160 : Conveyor;
  Conveyor70161 : Conveyor;
  Conveyor70162 : Conveyor;
  Conveyor70163 : Conveyor;
  Conveyor70164 : Conveyor;
  Conveyor70165 : Conveyor;
  Conveyor70166 : Conveyor;
  Conveyor70167 : Conveyor;
  Conveyor70168 : Conveyor;
  Conveyor70169 : Conveyor;
  Conveyor70170 : Conveyor;
  Conveyor70171 : Conveyor;
  Conveyor70172 : Conveyor;
  Conveyor70173 : Conveyor;
  Conveyor70174 : Conveyor;
  Conveyor70175 : Conveyor;
  Conveyor70176 : Conveyor;
  Conveyor70177 : Conveyor;
  Conveyor70178 : Conveyor;
  Conveyor70179 : Conveyor;
  Conveyor70180 : Conveyor;
  Conveyor70181 : Conveyor;
  Conveyor70182 : Conveyor;
  Conveyor70183 : Conveyor;
  Conveyor70184 : Conveyor;
  Conveyor70185 : Conveyor;
  Conveyor70186 : Conveyor;
  Conveyor70187 : Conveyor;
  Conveyor70188 : Conveyor;
  Conveyor70189 : Conveyor;
  Conveyor70190 : Conveyor;
  Conveyor70191 : Conveyor;
  Conveyor70192 : Conveyor;
  Conveyor70193 : Conveyor;
  Conveyor70194 : Conveyor;
  Conveyor70195 : Conveyor;
  Conveyor70196 : Conveyor;
  Conveyor70197 : Conveyor;
  Conveyor70198 : Conveyor;
  Conveyor70199 : Conveyor;
  Conveyor701100 : Conveyor;
  Conveyor701101 : Conveyor;
  Conveyor701102 : Conveyor;
  Conveyor701103 : Conveyor;
  Conveyor701104 : Conveyor;
  Conveyor701105 : Conveyor;
  Conveyor701106 : Conveyor;
  Conveyor701107 : Conveyor;
  Conveyor701108 : Conveyor;
  Conveyor701109 : Conveyor;
  Conveyor701110 : Conveyor;
  Conveyor701111 : Conveyor;
  Conveyor701112 : Conveyor;
  ConveyorIO70101 : ConveyorIO;
  ConveyorIO70102 : ConveyorIO;
  ConveyorIO70103 : ConveyorIO;
  ConveyorIO70104 : ConveyorIO;
  ConveyorIO70105 : ConveyorIO;
  ConveyorIO70106 : ConveyorIO;
  ConveyorIO70107 : ConveyorIO;
  ConveyorIO70108 : ConveyorIO;
  ConveyorIO70109 : ConveyorIO;
  ConveyorIO70110 : ConveyorIO;
  ConveyorIO70111 : ConveyorIO;
  ConveyorIO70112 : ConveyorIO;
  ConveyorIO70113 : ConveyorIO;
  ConveyorIO70114 : ConveyorIO;
  ConveyorIO70115 : ConveyorIO;
  ConveyorIO70116 : ConveyorIO;
  ConveyorIO70117 : ConveyorIO;
  ConveyorIO70118 : ConveyorIO;
  ConveyorIO70119 : ConveyorIO;
  ConveyorIO70120 : ConveyorIO;
  ConveyorIO70121 : ConveyorIO;
  ConveyorIO70122 : ConveyorIO;
  ConveyorIO70123 : ConveyorIO;
  ConveyorIO70124 : ConveyorIO;
  ConveyorIO70125 : ConveyorIO;
  ConveyorIO70126 : ConveyorIO;
  ConveyorIO70127 : ConveyorIO;
  ConveyorIO70128 : ConveyorIO;
  ConveyorIO70129 : ConveyorIO;
  ConveyorIO70130 : ConveyorIO;
  ConveyorIO70131 : ConveyorIO;
  ConveyorIO70132 : ConveyorIO;
  ConveyorIO70133 : ConveyorIO;
  ConveyorIO70134 : ConveyorIO;
  ConveyorIO70135 : ConveyorIO;
  ConveyorIO70136 : ConveyorIO;
  ConveyorIO70137 : ConveyorIO;
  ConveyorIO70138 : ConveyorIO;
  ConveyorIO70139 : ConveyorIO;
  ConveyorIO70140 : ConveyorIO;
  ConveyorIO70141 : ConveyorIO;
  ConveyorIO70142 : ConveyorIO;
  ConveyorIO70143 : ConveyorIO;
  ConveyorIO70144 : ConveyorIO;
  ConveyorIO70145 : ConveyorIO;
  ConveyorIO70146 : ConveyorIO;
  ConveyorIO70147 : ConveyorIO;
  ConveyorIO70148 : ConveyorIO;
  ConveyorIO70149 : ConveyorIO;
  ConveyorIO70150 : ConveyorIO;
  ConveyorIO70151 : ConveyorIO;
  ConveyorIO70152 : ConveyorIO;
  ConveyorIO70153 : ConveyorIO;
  ConveyorIO70154 : ConveyorIO;
  ConveyorIO70155 : ConveyorIO;
  ConveyorIO70156 : ConveyorIO;
  ConveyorIO70157 : ConveyorIO;
  ConveyorIO70158 : ConveyorIO;
  ConveyorIO70159 : ConveyorIO;
  ConveyorIO70160 : ConveyorIO;
  ConveyorIO70161 : ConveyorIO;
  ConveyorIO70162 : ConveyorIO;
  ConveyorIO70163 : ConveyorIO;
  ConveyorIO70164 : ConveyorIO;
  ConveyorIO70165 : ConveyorIO;
  ConveyorIO70166 : ConveyorIO;
  ConveyorIO70167 : ConveyorIO;
  ConveyorIO70168 : ConveyorIO;
  ConveyorIO70169 : ConveyorIO;
  ConveyorIO70170 : ConveyorIO;
  ConveyorIO70171 : ConveyorIO;
  ConveyorIO70172 : ConveyorIO;
  ConveyorIO70173 : ConveyorIO;
  ConveyorIO70174 : ConveyorIO;
  ConveyorIO70175 : ConveyorIO;
  ConveyorIO70176 : ConveyorIO;
  ConveyorIO70177 : ConveyorIO;
  ConveyorIO70178 : ConveyorIO;
  ConveyorIO70179 : ConveyorIO;
  ConveyorIO70180 : ConveyorIO;
  ConveyorIO70181 : ConveyorIO;
  ConveyorIO70182 : ConveyorIO;
  ConveyorIO70183 : ConveyorIO;
  ConveyorIO70184 : ConveyorIO;
  ConveyorIO70185 : ConveyorIO;
  ConveyorIO70186 : ConveyorIO;
  ConveyorIO70187 : ConveyorIO;
  ConveyorIO70188 : ConveyorIO;
  ConveyorIO70189 : ConveyorIO;
  ConveyorIO70190 : ConveyorIO;
  ConveyorIO70191 : ConveyorIO;
  ConveyorIO70192 : ConveyorIO;
  ConveyorIO70193 : ConveyorIO;
  ConveyorIO70194 : ConveyorIO;
  ConveyorIO70195 : ConveyorIO;
  ConveyorIO70196 : ConveyorIO;
  ConveyorIO70197 : ConveyorIO;
  ConveyorIO70198 : ConveyorIO;
  ConveyorIO70199 : ConveyorIO;
  ConveyorIO701100 : ConveyorIO;